 986 '~S001R11 Sealer Ctrlr 2 Required Rezeroing WB2[30].26'; 987 '~S001R11 Mig Barrel Replacement Warning WB2[30].27'; 988 '~S001R11 Mig Barrel Replacement Required WB2[30].28'; 989 '~S001R11 In Touch Up Mode WB2[30].29'; 990 '~S001R11 Touch Up Mode Not Enabled WB2[30].30'; 991 '~Spare WB2[30].31'; 992 '~S001R11 Laser Controller Fault WB2[31].0'; 993 '~S001R11 Laser Dirty Glass Warning WB2[31].1'; 994 '~S001R11 Laser Warning WB2[31].2'; 995 '~Spare WB2[31].3'; 996 '~Spare WB2[31].4'; 997 '~Spare WB2[31].5'; 998 '~Spare WB2[31].6'; 999 '~Spare WB2[31].7'; 1000 '~Spare WB2[31].8'; 1001 '~Spare WB2[31].9'; 1002 '~Spare WB2[31].10'; 1003 '~Spare WB2[31].11'; 1004 '~Spare WB2[31].12'; 1005 '~Spare WB2[31].13'; 1006 '~Spare WB2[31].14'; 1007 '~Spare WB2[31].15'; 1008 '~Spare WB2[31].16'; 1009 '~Spare WB2[31].17'; 1010 '~Spare WB2[31].18'; 1011 '~Spare WB2[31].19'; 1012 '~Spare WB2[31].20'; 1013 '~Spare WB2[31].21'; 1014 '~Spare WB2[31].22'; 1015 '~Spare WB2[31].23'; 1016 '~Spare WB2[31].24'; 1017 '~Spare WB2[31].25'; 1018 '~Spare WB2[31].26'; 1019 '~Spare WB2[31].27'; 1020 '~Spare WB2[31].28'; 1021 '~Spare WB2[31].29'; 1022 '~Spare WB2[31].30'; 1023 '~Spare WB2[31].31'; 1024 '~Spare WB2[32].0'; 1025 '~Spare WB2[32].1'; 1026 '~Spare WB2[32].2'; 1027 '~Spare WB2[32].3'; 1028 '~Spare WB2[32].4'; 1029 '~Spare WB2[32].5'; 1030 '~Spare WB2[32].6'; 1031 '~Spare WB2[32].7'; 1032 '~Spare WB2[32].8'; 1033 '~Spare WB2[32].9'; 1034 '~Spare WB2[32].10'; 1035 '~Spare WB2[32].11'; 1036 '~Spare WB2[32].12'; 1037 '~Spare WB2[32].13'; 1038 '~Spare WB2[32].14'; 1039 '~Spare WB2[32].15'; 1040 '~Spare WB2[32].16'; 1041 '~Spare WB2[32].17'; 1042 '~Spare WB2[32].18'; 1043 '~Spare WB2[32].19'; 1044 '~Spare WB2[32].20'; 1045 '~Spare WB2[32].21'; 1046 '~Spare WB2[32].22'; 1047 '~Spare WB2[32].23'; 1048 '~Spare WB2[32].24'; 1049 '~Spare WB2[32].25'; 1050 '~Spare WB2[32].26'; 1051 '~Spare WB2[32].27'; 1052 '~Spare WB2[32].28'; 1053 '~Spare WB2[32].29'; 1054 '~Spare WB2[32].30'; 1055 '~Spare WB2[32].31'; 1056 '~Spare WB2[33].0'; 1057 '~Spare WB2[33].1'; 1058 '~Spare WB2[33].2'; 1059 '~Spare WB2[33].3'; 1060 '~Spare WB2[33].4'; 1061 '~Spare WB2[33].5'; 1062 '~Spare WB2[33].6'; 1063 '~Spare WB2[33].7'; 1064 '~Spare WB2[33].8'; 1065 '~Spare WB2[33].9'; 1066 '~Spare WB2[33].10'; 1067 '~Spare WB2[33].11'; 1068 '~Spare WB2[33].12'; 1069 '~Spare WB2[33].13'; 1070 '~Spare WB2[33].14'; 1071 '~Spare WB2[33].15'; 1072 '~Spare WB2[33].16'; 1073 '~Spare WB2[33].17'; 1074 '~Spare WB2[33].18'; 1075 '~Spare WB2[33].19'; 1076 '~Spare WB2[33].20'; 1077 '~Spare WB2[33].21'; 1078 '~Spare WB2[33].22'; 1079 '~Spare WB2[33].23'; 1080 '~Spare WB2[33].24'; 1081 '~Spare WB2[33].25'; 1082 '~Spare WB2[33].26'; 1083 '~Spare WB2[33].27'; 1084 '~Spare WB2[33].28'; 1085 '~Spare WB2[33].29'; 1086 '~Spare WB2[33].30'; 1087 '~Spare WB2[33].31'; 1088 '~S001R12 Waiting Zone #1 Not Clear WB2[34].0'; 1089 '~S001R12 Waiting Zone #2 Not Clear WB2[34].1'; 1090 '~S001R12 Waiting Zone #3 Not Clear WB2[34].2'; 1091 '~S001R12 Waiting Zone #4 Not Clear WB2[34].3'; 1092 '~S001R12 Waiting Zone #5 Not Clear WB2[34].4'; 1093 '~S001R12 Waiting Zone #6 Not Clear WB2[34].5'; 1094 '~S001R12 Waiting Zone #7 Not Clear WB2[34].6'; 1095 '~S001R12 Waiting Zone #8 Not Clear WB2[34].7'; 1096 '~S001R12 Waiting Zone #9 Not Clear WB2[34].8'; 1097 '~S001R12 Waiting Zone #10 Not Clear WB2[34].9'; 1098 '~S001R12 Waiting Zone #11 Not Clear WB2[34].10'; 1099 '~S001R12 Waiting Zone #12 Not Clear WB2[34].11'; 1100 '~S001R12 Waiting Zone #13 Not Clear WB2[34].12'; 1101 '~S001R12 Waiting Zone #14 Not Clear WB2[34].13'; 1102 '~S001R12 Waiting Tip Dress Zone #1 Not Clear WB2[34].14'; 1103 '~S001R12 Waiting Tip Dress Zone #2 Not Clear WB2[34].15'; 1104 '~S001R12 Adjacent Robot xx-xx In Teach WB2[34].16'; 1105 '~S001R12 Adjacent Robot xx-xx In Teach WB2[34].17'; 1106 '~S001R12 Adjacent Robot xx-xx In Teach WB2[34].18'; 1107 '~S001R12 Adjacent Robot xx-xx In Teach WB2[34].19'; 1108 '~S001R12 Adjacent Robot xx-xx In Teach WB2[34].20'; 1109 '~S001R12 Adjacent Robot xx-xx In Teach WB2[34].21'; 1110 '~S001R12 Adjacent Robot xx-xx In Teach WB2[34].22'; 1111 '~S001R12 Adjacent Robot xx-xx In Teach WB2[34].23'; 1112 '~S001R12 Adjacent Robot xx-xx In Teach WB2[34].24'; 1113 '~S001R12 Adjacent Robot xx-xx In Teach WB2[34].25'; 1114 '~Spare WB2[34].26'; 1115 '~Spare WB2[34].27'; 1116 '~Spare WB2[34].28'; 1117 '~S001R12 Robot Not Clear Of Fixture WB2[34].29'; 1118 '~Spare WB2[34].30'; 1119 '~Spare WB2[34].31'; 1120 '~Spare WB2[35].0'; 1121 '~Spare WB2[35].1'; 1122 '~Spare WB2[35].2'; 1123 '~Spare WB2[35].3'; 1124 '~Spare WB2[35].4'; 1125 '~Spare WB2[35].5'; 1126 '~Spare WB2[35].6'; 1127 '~Spare WB2[35].7'; 1128 '~Spare WB2[35].8'; 1129 '~Spare WB2[35].9'; 1130 '~Spare WB2[35].10'; 1131 '~Spare WB2[35].11'; 1132 '~Spare WB2[35].12'; 1133 '~Spare WB2[35].13'; 1134 '~Spare WB2[35].14'; 1135 '~Spare WB2[35].15'; 1136 '~Spare WB2[35].16'; 1137 '~Spare WB2[35].17'; 1138 '~Spare WB2[35].18'; 1139 '~Spare WB2[35].19'; 1140 '~Spare WB2[35].20'; 1141 '~Spare WB2[35].21'; 1142 '~Spare WB2[35].22'; 1143 '~Spare WB2[35].23'; 1144 '~Spare WB2[35].24'; 1145 '~Spare WB2[35].25'; 1146 '~Spare WB2[35].26'; 1147 '~Spare WB2[35].27'; 1148 '~Spare WB2[35].28'; 1149 '~Spare WB2[35].29'; 1150 '~Spare WB2[35].30'; 1151 '~Spare WB2[35].31'; 1152 '~S001R12 Cycle Overtime WB2[36].0'; 1153 '~S001R12 In Bypass WB2[36].1'; 1154 '~S001R12 Battery Low WB2[36].2'; 1155 '~S001R12 Servo Over Torque WB2[36].3'; 1156 '~S001R12 Process Retry In Progress WB2[36].4'; 1157 '~Spare WB2[36].5'; 1158 '~S001R12 Robot Edit Occurred Ext App WB2[36].6'; 1159 '~S001R12 Robot Input Simmed WB2[36].7'; 1160 '~S001R12 Robot Output Simmed WB2[36].8'; 1161 '~Spare WB2[36].9'; 1162 '~Spare WB2[36].10'; 1163 '~Spare WB2[36].11'; 1164 '~Spare WB2[36].12'; 1165 '~Spare WB2[36].13'; 1166 '~Spare WB2[36].14'; 1167 '~Spare WB2[36].15'; 1168 '~S001R12F1B1.M.ModuleFlt - Externa App 1 I/O Module Warning WB2[36].16'; 1169 '~S001R12F2B1.M.ModuleFlt - Externa App 2 I/O Module Warning WB2[36].17'; 1170 '~S001R12F3B1.M.ModuleFlt - Externa App 3 I/O Module Warning WB2[36].18'; 1171 '~Spare WB2[36].19'; 1172 '~Spare WB2[36].20'; 1173 '~Spare WB2[36].21'; 1174 '~Spare WB2[36].22'; 1175 '~Spare WB2[36].23'; 1176 '~S001R12ES1 - S001R12 EtherNet Switch Port At Half Duplex WB2[36].24'; 1177 '~S001R12ES1 - S001R12 EtherNet Switch Config Changes Not Saved WB2[36].25'; 1178 '~S001R12ES1 - S001R12 EtherNet Switch Configuration Changed WB2[36].26'; 1179 '~S001R12ES1 - S001R12 EtherNet Switch Port With Excessive Errors WB2[36].27'; 1180 '~S001R12ES1 - S001R12 EtherNet Switch Port With Utilization Warning WB2[36].28'; 1181 '~S001R12ES1 - S001R12 EtherNet Switch Changes Require Reboot WB2[36].29'; 1182 '~Spare WB2[36].30'; 1183 '~Spare WB2[36].31'; 1184 '~Spare WB2[37].0'; 1185 '~Spare WB2[37].1'; 1186 '~S001R12 Servo Gun Tip Calib Request 1 WB2[37].2'; 1187 '~S001R12 I-Available Warning 1 WB2[37].3'; 1188 '~S001R12 Tip Dress Motor 1 Fault Bypassed WB2[37].4'; 1189 '~S001R12 Tip Change Notice 1 WB2[37].5'; 1190 '~S001R12 Bypass Tip Dresser 1 Selected WB2[37].6'; 1191 '~S001R12 Auto Tip Changer Low 1 WB2[37].7'; 1192 '~S001R12 Auto Tip Changer Empty 1 WB2[37].8'; 1193 '~S001R12 Tip Wear Ratio Warning 1 - Touch Up Tip Dress Program WB2[37].9'; 1194 '~S001R12 Stud Weld 1 Maintenance Reqd WB2[37].10'; 1195 '~S001R12 Stud Weld 1 Low Stud Warning WB2[37].11'; 1196 '~Spare WB2[37].12'; 1197 '~S001R12 Rivet 1 Low Rivet Warning WB2[37].13'; 1198 '~S001R12 Rivet 1 - Skip Once Initiated from Robot TP WB2[37].14'; 1199 '~S001R12 Rivet 1 - Skip Remaining Initiated from Robot TP WB2[37].15'; 1200 '~S001R12 Rivet 1 Preventive Maintenace Required WB2[37].16'; 1201 '~S001R12 Rivet 1 Magazine Low WB2[37].17'; 1202 '~S001R12 Tip Change 1 Bypassed WB2[37].18'; 1203 '~S001R12 Mig Weld Fluid Level Low WB2[37].19'; 1204 '~S001R12 Weld Ctrlr 1 Adaptive Mode Is Disabled WB2[37].20'; 1205 '~S001R12 Tip Cutter 1 Warning WB2[37].21'; 1206 '~S001R12 Rivet 1 Tape-Cut Required WB2[37].22'; 1207 '~S001R12 Wire Feeder Motor Over Current WB2[37].23'; 1208 '~Spare WB2[37].24'; 1209 '~S001R12 Sealer Ctrlr 1 Minor Fault WB2[37].25'; 1210 '~S001R12 Sealer Ctrlr 1 Required Rezeroing WB2[37].26'; 1211 '~S001R12 Loaded To Average WB2[37].27'; 1212 '~S001R12 Vision Process Aborted WB2[37].28'; 1213 '~S001R12 Vision System Trending WB2[37].29'; 1214 '~S001R12 Vision Out Of Tolerance WB2[37].30'; 1215 '~Spare WB2[37].31'; 1216 '~Spare WB2[38].0'; 1217 '~Spare WB2[38].1'; 1218 '~S001R12 Servo Gun Tip Calib Request 2 WB2[38].2'; 1219 '~S001R12 I-Available Warning 2 WB2[38].3'; 1220 '~S001R12 Tip Dress Motor 2 Fault Bypassed WB2[38].4'; 1221 '~S001R12 Tip Change Notice 2 WB2[38].5'; 1222 '~S001R12 Bypass Tip Dresser 2 Selected WB2[38].6'; 1223 '~S001R12 Auto Tip Changer Low 2 WB2[38].7'; 1224 '~S001R12 Auto Tip Changer Empty 2 WB2[38].8'; 1225 '~S001R12 Tip Wear Ratio Warning 2 - Touch Up Tip Dress Program WB2[38].9'; 1226 '~S001R12 Stud Weld 2 Maintenance Reqd WB2[38].10'; 1227 '~S001R12 Stud Weld 2 Low Stud Warning WB2[38].11'; 1228 '~Spare WB2[38].12'; 1229 '~S001R12 Rivet 2 Low Rivet Warning WB2[38].13'; 1230 '~S001R12 Rivet 2 - Skip Once Initiated from Robot TP WB2[38].14'; 1231 '~S001R12 Rivet 2 - Skip Remaining Initiated from Robot TP WB2[38].15'; 1232 '~S001R12 Rivet 2 Preventive Maintenace Required WB2[38].16'; 1233 '~S001R12 Rivet 2 Magazine Low WB2[38].17'; 1234 '~S001R12 Tip Change 2 Bypassed WB2[38].18'; 1235 '~S001R12 Laser Dirty Glass Warning WB2[38].19'; 1236 '~S001R12 Weld Ctrlr 2 Adaptive Mode Is Disabled WB2[38].20'; 1237 '~S001R12 Tip Cutter 2 Warning WB2[38].21'; 1238 '~S001R12 Rivet 2 Tape-Cut Required WB2[38].22'; 1239 '~S001R12 Mig Tip Nozzel Replacement Warning WB2[38].23'; 1240 '~S001R12 Mig Tip Nozzel Replacement Required WB2[38].24'; 1241 '~S001R12 Sealer Ctrlr 2 Minor Fault WB2[38].25'; 1242 '~S001R12 Sealer Ctrlr 2 Required Rezeroing WB2[38].26'; 1243 '~S001R12 Mig Barrel Replacement Warning WB2[38].27'; 1244 '~S001R12 Mig Barrel Replacement Required WB2[38].28'; 1245 '~S001R12 In Touch Up Mode WB2[38].29'; 1246 '~S001R12 Touch Up Mode Not Enabled WB2[38].30'; 1247 '~Spare WB2[38].31'; 1248 '~S001R12 Laser Controller Fault WB2[39].0'; 1249 '~S001R12 Laser Dirty Glass Warning WB2[39].1'; 1250 '~S001R12 Laser Warning WB2[39].2'; 1251 '~Spare WB2[39].3'; 1252 '~Spare WB2[39].4'; 1253 '~Spare WB2[39].5'; 1254 '~Spare WB2[39].6'; 1255 '~Spare WB2[39].7'; 1256 '~Spare WB2[39].8'; 1257 '~Spare WB2[39].9'; 1258 '~Spare WB2[39].10'; 1259 '~Spare WB2[39].11'; 1260 '~Spare WB2[39].12'; 1261 '~Spare WB2[39].13'; 1262 '~Spare WB2[39].14'; 1263 '~Spare WB2[39].15'; 1264 '~Spare WB2[39].16'; 1265 '~Spare WB2[39].17'; 1266 '~Spare WB2[39].18'; 1267 '~Spare WB2[39].19'; 1268 '~Spare WB2[39].20'; 1269 '~Spare WB2[39].21'; 1270 '~Spare WB2[39].22'; 1271 '~Spare WB2[39].23'; 1272 '~Spare WB2[39].24'; 1273 '~Spare WB2[39].25'; 1274 '~Spare WB2[39].26'; 1275 '~Spare WB2[39].27'; 1276 '~Spare WB2[39].28'; 1277 '~Spare WB2[39].29'; 1278 '~Spare WB2[39].30'; 1279 '~Spare WB2[39].31'; 1280 '~Spare WB2[40].0'; 1281 '~Spare WB2[40].1'; 1282 '~Spare WB2[40].2'; 1283 '~Spare WB2[40].3'; 1284 '~Spare WB2[40].4'; 1285 '~Spare WB2[40].5'; 1286 '~Spare WB2[40].6'; 1287 '~Spare WB2[40].7'; 1288 '~Spare WB2[40].8'; 1289 '~Spare WB2[40].9'; 1290 '~Spare WB2[40].10'; 1291 '~Spare WB2[40].11'; 1292 '~Spare WB2[40].12'; 1293 '~Spare WB2[40].13'; 1294 '~Spare WB2[40].14'; 1295 '~Spare WB2[40].15'; 1296 '~Spare WB2[40].16'; 1297 '~Spare WB2[40].17'; 1298 '~Spare WB2[40].18'; 1299 '~Spare WB2[40].19'; 1300 '~Spare WB2[40].20'; 1301 '~Spare WB2[40].21'; 1302 '~Spare WB2[40].22'; 1303 '~Spare WB2[40].23'; 1304 '~Spare WB2[40].24'; 1305 '~Spare WB2[40].25'; 1306 '~Spare WB2[40].26'; 1307 '~Spare WB2[40].27'; 1308 '~Spare WB2[40].28'; 1309 '~Spare WB2[40].29'; 1310 '~Spare WB2[40].30'; 1311 '~Spare WB2[40].31'; 1312 '~Spare WB2[41].0'; 1313 '~Spare WB2[41].1'; 1314 '~Spare WB2[41].2'; 1315 '~Spare WB2[41].3'; 1316 '~Spare WB2[41].4'; 1317 '~Spare WB2[41].5'; 1318 '~Spare WB2[41].6'; 1319 '~Spare WB2[41].7'; 1320 '~Spare WB2[41].8'; 1321 '~Spare WB2[41].9'; 1322 '~Spare WB2[41].10'; 1323 '~Spare WB2[41].11'; 1324 '~Spare WB2[41].12'; 1325 '~Spare WB2[41].13'; 1326 '~Spare WB2[41].14'; 1327 '~Spare WB2[41].15'; 1328 '~Spare WB2[41].16'; 1329 '~Spare WB2[41].17'; 1330 '~Spare WB2[41].18'; 1331 '~Spare WB2[41].19'; 1332 '~Spare WB2[41].20'; 1333 '~Spare WB2[41].21'; 1334 '~Spare WB2[41].22'; 1335 '~Spare WB2[41].23'; 1336 '~Spare WB2[41].24'; 1337 '~Spare WB2[41].25'; 1338 '~Spare WB2[41].26'; 1339 '~Spare WB2[41].27'; 1340 '~Spare WB2[41].28'; 1341 '~Spare WB2[41].29'; 1342 '~Spare WB2[41].30'; 1343 '~Spare WB2[41].31'; 1344 '~S001R13 Waiting Zone #1 Not Clear WB2[42].0'; 1345 '~S001R13 Waiting Zone #2 Not Clear WB2[42].1'; 1346 '~S001R13 Waiting Zone #3 Not Clear WB2[42].2'; 1347 '~S001R13 Waiting Zone #4 Not Clear WB2[42].3'; 1348 '~S001R13 Waiting Zone #5 Not Clear WB2[42].4'; 1349 '~S001R13 Waiting Zone #6 Not Clear WB2[42].5'; 1350 '~S001R13 Waiting Zone #7 Not Clear WB2[42].6'; 1351 '~S001R13 Waiting Zone #8 Not Clear WB2[42].7'; 1352 '~S001R13 Waiting Zone #9 Not Clear WB2[42].8'; 1353 '~S001R13 Waiting Zone #10 Not Clear WB2[42].9'; 1354 '~S001R13 Waiting Zone #11 Not Clear WB2[42].10'; 1355 '~S001R13 Waiting Zone #12 Not Clear WB2[42].11'; 1356 '~S001R13 Waiting Zone #13 Not Clear WB2[42].12'; 1357 '~S001R13 Waiting Zone #14 Not Clear WB2[42].13'; 1358 '~S001R13 Waiting Tip Dress Zone #1 Not Clear WB2[42].14'; 1359 '~S001R13 Waiting Tip Dress Zone #2 Not Clear WB2[42].15'; 1360 '~S001R13 Adjacent Robot xx-xx In Teach WB2[42].16'; 1361 '~S001R13 Adjacent Robot xx-xx In Teach WB2[42].17'; 1362 '~S001R13 Adjacent Robot xx-xx In Teach WB2[42].18'; 1363 '~S001R13 Adjacent Robot xx-xx In Teach WB2[42].19'; 1364 '~S001R13 Adjacent Robot xx-xx In Teach WB2[42].20'; 1365 '~S001R13 Adjacent Robot xx-xx In Teach WB2[42].21'; 1366 '~S001R13 Adjacent Robot xx-xx In Teach WB2[42].22'; 1367 '~S001R13 Adjacent Robot xx-xx In Teach WB2[42].23'; 1368 '~S001R13 Adjacent Robot xx-xx In Teach WB2[42].24'; 1369 '~S001R13 Adjacent Robot xx-xx In Teach WB2[42].25'; 1370 '~Spare WB2[42].26'; 1371 '~Spare WB2[42].27'; 1372 '~Spare WB2[42].28'; 1373 '~S001R13 Robot Not Clear Of Fixture WB2[42].29'; 1374 '~Spare WB2[42].30'; 1375 '~Spare WB2[42].31'; 1376 '~Spare WB2[43].0'; 1377 '~Spare WB2[43].1'; 1378 '~Spare WB2[43].2'; 1379 '~Spare WB2[43].3'; 1380 '~Spare WB2[43].4'; 1381 '~Spare WB2[43].5'; 1382 '~Spare WB2[43].6'; 1383 '~Spare WB2[43].7'; 1384 '~Spare WB2[43].8'; 1385 '~Spare WB2[43].9'; 1386 '~Spare WB2[43].10'; 1387 '~Spare WB2[43].11'; 1388 '~Spare WB2[43].12'; 1389 '~Spare WB2[43].13'; 1390 '~Spare WB2[43].14'; 1391 '~Spare WB2[43].15'; 1392 '~Spare WB2[43].16'; 1393 '~Spare WB2[43].17'; 1394 '~Spare WB2[43].18'; 1395 '~Spare WB2[43].19'; 1396 '~Spare WB2[43].20'; 1397 '~Spare WB2[43].21'; 1398 '~Spare WB2[43].22'; 1399 '~Spare WB2[43].23'; 1400 '~Spare WB2[43].24'; 1401 '~Spare WB2[43].25'; 1402 '~Spare WB2[43].26'; 1403 '~Spare WB2[43].27'; 1404 '~Spare WB2[43].28'; 1405 '~Spare WB2[43].29'; 1406 '~Spare WB2[43].30'; 1407 '~Spare WB2[43].31'; 1408 '~S001R13 Cycle Overtime WB2[44].0'; 1409 '~S001R13 In Bypass WB2[44].1'; 1410 '~S001R13 Battery Low WB2[44].2'; 1411 '~S001R13 Servo Over Torque WB2[44].3'; 1412 '~S001R13 Process Retry In Progress WB2[44].4'; 1413 '~Spare WB2[44].5'; 1414 '~S001R13 Robot Edit Occurred Ext App WB2[44].6'; 1415 '~S001R13 Robot Input Simmed WB2[44].7'; 1416 '~S001R13 Robot Output Simmed WB2[44].8'; 1417 '~Spare WB2[44].9'; 1418 '~Spare WB2[44].10'; 1419 '~Spare WB2[44].11'; 1420 '~Spare WB2[44].12'; 1421 '~Spare WB2[44].13'; 1422 '~Spare WB2[44].14'; 1423 '~Spare WB2[44].15'; 1424 '~S001R13F1B1.M.ModuleFlt - Externa App 1 I/O Module Warning WB2[44].16'; 1425 '~S001R13F2B1.M.ModuleFlt - Externa App 2 I/O Module Warning WB2[44].17'; 1426 '~S001R13F3B1.M.ModuleFlt - Externa App 3 I/O Module Warning WB2[44].18'; 1427 '~Spare WB2[44].19'; 1428 '~Spare WB2[44].20'; 1429 '~Spare WB2[44].21'; 1430 '~Spare WB2[44].22'; 1431 '~Spare WB2[44].23'; 1432 '~S001R13ES1 - S001R13 EtherNet Switch Port At Half Duplex WB2[44].24'; 1433 '~S001R13ES1 - S001R13 EtherNet Switch Config Changes Not Saved WB2[44].25'; 1434 '~S001R13ES1 - S001R13 EtherNet Switch Configuration Changed WB2[44].26'; 1435 '~S001R13ES1 - S001R13 EtherNet Switch Port With Excessive Errors WB2[44].27'; 1436 '~S001R13ES1 - S001R13 EtherNet Switch Port With Utilization Warning WB2[44].28'; 1437 '~S001R13ES1 - S001R13 EtherNet Switch Changes Require Reboot WB2[44].29'; 1438 '~Spare WB2[44].30'; 1439 '~Spare WB2[44].31'; 1440 '~Spare WB2[45].0'; 1441 '~Spare WB2[45].1'; 1442 '~S001R13 Servo Gun Tip Calib Request 1 WB2[45].2'; 1443 '~S001R13 I-Available Warning 1 WB2[45].3'; 1444 '~S001R13 Tip Dress Motor 1 Fault Bypassed WB2[45].4'; 1445 '~S001R13 Tip Change Notice 1 WB2[45].5'; 1446 '~S001R13 Bypass Tip Dresser 1 Selected WB2[45].6'; 1447 '~S001R13 Auto Tip Changer Low 1 WB2[45].7'; 1448 '~S001R13 Auto Tip Changer Empty 1 WB2[45].8'; 1449 '~S001R13 Tip Wear Ratio Warning 1 - Touch Up Tip Dress Program WB2[45].9'; 1450 '~S001R13 Stud Weld 1 Maintenance Reqd WB2[45].10'; 1451 '~S001R13 Stud Weld 1 Low Stud Warning WB2[45].11'; 1452 '~Spare WB2[45].12'; 1453 '~S001R13 Rivet 1 Low Rivet Warning WB2[45].13'; 1454 '~S001R13 Rivet 1 - Skip Once Initiated from Robot TP WB2[45].14'; 1455 '~S001R13 Rivet 1 - Skip Remaining Initiated from Robot TP WB2[45].15'; 1456 '~S001R13 Rivet 1 Preventive Maintenace Required WB2[45].16'; 1457 '~S001R13 Rivet 1 Magazine Low WB2[45].17'; 1458 '~S001R13 Tip Change 1 Bypassed WB2[45].18'; 1459 '~S001R13 Mig Weld Fluid Level Low WB2[45].19'; 1460 '~S001R13 Weld Ctrlr 1 Adaptive Mode Is Disabled WB2[45].20'; 1461 '~S001R13 Tip Cutter 1 Warning WB2[45].21'; 1462 '~S001R13 Rivet 1 Tape-Cut Required WB2[45].22'; 1463 '~S001R13 Wire Feeder Motor Over Current WB2[45].23'; 1464 '~Spare WB2[45].24'; 1465 '~S001R13 Sealer Ctrlr 1 Minor Fault WB2[45].25'; 1466 '~S001R13 Sealer Ctrlr 1 Required Rezeroing WB2[45].26'; 1467 '~S001R13 Loaded To Average WB2[45].27'; 1468 '~S001R13 Vision Process Aborted WB2[45].28'; 1469 '~S001R13 Vision System Trending WB2[45].29'; 1470 '~S001R13 Vision Out Of Tolerance WB2[45].30'; 1471 '~Spare WB2[45].31'; 1472 '~Spare WB2[46].0'; 1473 '~Spare WB2[46].1'; 1474 '~S001R13 Servo Gun Tip Calib Request 2 WB2[46].2'; 1475 '~S001R13 I-Available Warning 2 WB2[46].3'; 1476 '~S001R13 Tip Dress Motor 2 Fault Bypassed WB2[46].4'; 1477 '~S001R13 Tip Change Notice 2 WB2[46].5'; 1478 '~S001R13 Bypass Tip Dresser 2 Selected WB2[46].6'; 1479 '~S001R13 Auto Tip Changer Low 2 WB2[46].7'; 1480 '~S001R13 Auto Tip Changer Empty 2 WB2[46].8'; 1481 '~S001R13 Tip Wear Ratio Warning 2 - Touch Up Tip Dress Program WB2[46].9'; 1482 '~S001R13 Stud Weld 2 Maintenance Reqd WB2[46].10'; 1483 '~S001R13 Stud Weld 2 Low Stud Warning WB2[46].11'; 1484 '~Spare WB2[46].12'; 1485 '~S001R13 Rivet 2 Low Rivet Warning WB2[46].13'; 1486 '~S001R13 Rivet 2 - Skip Once Initiated from Robot TP WB2[46].14'; 1487 '~S001R13 Rivet 2 - Skip Remaining Initiated from Robot TP WB2[46].15'; 1488 '~S001R13 Rivet 2 Preventive Maintenace Required WB2[46].16'; 1489 '~S001R13 Rivet 2 Magazine Low WB2[46].17'; 1490 '~S001R13 Tip Change 2 Bypassed WB2[46].18'; 1491 '~S001R13 Laser Dirty Glass Warning WB2[46].19'; 1492 '~S001R13 Weld Ctrlr 2 Adaptive Mode Is Disabled WB2[46].20'; 1493 '~S001R13 Tip Cutter 2 Warning WB2[46].21'; 1494 '~S001R13 Rivet 2 Tape-Cut Required WB2[46].22'; 1495 '~S001R13 Mig Tip Nozzel Replacement Warning WB2[46].23'; 1496 '~S001R13 Mig Tip Nozzel Replacement Required WB2[46].24'; 1497 '~S001R13 Sealer Ctrlr 2 Minor Fault WB2[46].25'; 1498 '~S001R13 Sealer Ctrlr 2 Required Rezeroing WB2[46].26'; 1499 '~S001R13 Mig Barrel Replacement Warning WB2[46].27'; 1500 '~S001R13 Mig Barrel Replacement Required WB2[46].28'; 1501 '~S001R13 In Touch Up Mode WB2[46].29'; 1502 '~S001R13 Touch Up Mode Not Enabled WB2[46].30'; 1503 '~Spare WB2[46].31'; 1504 '~S001R13 Laser Controller Fault WB2[47].0'; 1505 '~S001R13 Laser Dirty Glass Warning WB2[47].1'; 1506 '~S001R13 Laser Warning WB2[47].2'; 1507 '~Spare WB2[47].3'; 1508 '~Spare WB2[47].4'; 1509 '~Spare WB2[47].5'; 1510 '~Spare WB2[47].6'; 1511 '~Spare WB2[47].7'; 1512 '~Spare WB2[47].8'; 1513 '~Spare WB2[47].9'; 1514 '~Spare WB2[47].10'; 1515 '~Spare WB2[47].11'; 1516 '~Spare WB2[47].12'; 1517 '~Spare WB2[47].13'; 1518 '~Spare WB2[47].14'; 1519 '~Spare WB2[47].15'; 1520 '~Spare WB2[47].16'; 1521 '~Spare WB2[47].17'; 1522 '~Spare WB2[47].18'; 1523 '~Spare WB2[47].19'; 1524 '~Spare WB2[47].20'; 1525 '~Spare WB2[47].21'; 1526 '~Spare WB2[47].22'; 1527 '~Spare WB2[47].23'; 1528 '~Spare WB2[47].24'; 1529 '~Spare WB2[47].25'; 1530 '~Spare WB2[47].26'; 1531 '~Spare WB2[47].27'; 1532 '~Spare WB2[47].28'; 1533 '~Spare WB2[47].29'; 1534 '~Spare WB2[47].30'; 1535 '~Spare WB2[47].31'; 1536 '~Spare WB2[48].0'; 1537 '~Spare WB2[48].1'; 1538 '~Spare WB2[48].2'; 1539 '~Spare WB2[48].3'; 1540 '~Spare WB2[48].4'; 1541 '~Spare WB2[48].5'; 1542 '~Spare WB2[48].6'; 1543 '~Spare WB2[48].7'; 1544 '~Spare WB2[48].8'; 1545 '~Spare WB2[48].9'; 1546 '~Spare WB2[48].10'; 1547 '~Spare WB2[48].11'; 1548 '~Spare WB2[48].12'; 1549 '~Spare WB2[48].13'; 1550 '~Spare WB2[48].14'; 1551 '~Spare WB2[48].15'; 1552 '~Spare WB2[48].16'; 1553 '~Spare WB2[48].17'; 1554 '~Spare WB2[48].18'; 1555 '~Spare WB2[48].19'; 1556 '~Spare WB2[48].20'; 1557 '~Spare WB2[48].21'; 1558 '~Spare WB2[48].22'; 1559 '~Spare WB2[48].23'; 1560 '~Spare WB2[48].24'; 1561 '~Spare WB2[48].25'; 1562 '~Spare WB2[48].26'; 1563 '~Spare WB2[48].27'; 1564 '~Spare WB2[48].28'; 1565 '~Spare WB2[48].29'; 1566 '~Spare WB2[48].30'; 1567 '~Spare WB2[48].31'; 1568 '~Spare WB2[49].0'; 1569 '~Spare WB2[49].1'; 1570 '~Spare WB2[49].2'; 1571 '~Spare WB2[49].3'; 1572 '~Spare WB2[49].4'; 1573 '~Spare WB2[49].5'; 1574 '~Spare WB2[49].6'; 1575 '~Spare WB2[49].7'; 1576 '~Spare WB2[49].8'; 1577 '~Spare WB2[49].9'; 1578 '~Spare WB2[49].10'; 1579 '~Spare WB2[49].11'; 1580 '~Spare WB2[49].12'; 1581 '~Spare WB2[49].13'; 1582 '~Spare WB2[49].14'; 1583 '~Spare WB2[49].15'; 1584 '~Spare WB2[49].16'; 1585 '~Spare WB2[49].17'; 1586 '~Spare WB2[49].18'; 1587 '~Spare WB2[49].19'; 1588 '~Spare WB2[49].20'; 1589 '~Spare WB2[49].21'; 1590 '~Spare WB2[49].22'; 1591 '~Spare WB2[49].23'; 1592 '~Spare WB2[49].24'; 1593 '~Spare WB2[49].25'; 1594 '~Spare WB2[49].26'; 1595 '~Spare WB2[49].27'; 1596 '~Spare WB2[49].28'; 1597 '~Spare WB2[49].29'; 1598 '~Spare WB2[49].30'; 1599 '~Spare WB2[49].31'; 1600 '~S001R14 Waiting Zone #1 Not Clear WB2[50].0'; 1601 '~S001R14 Waiting Zone #2 Not Clear WB2[50].1'; 1602 '~S001R14 Waiting Zone #3 Not Clear WB2[50].2'; 1603 '~S001R14 Waiting Zone #4 Not Clear WB2[50].3'; 1604 '~S001R14 Waiting Zone #5 Not Clear WB2[50].4'; 1605 '~S001R14 Waiting Zone #6 Not Clear WB2[50].5'; 1606 '~S001R14 Waiting Zone #7 Not Clear WB2[50].6'; 1607 '~S001R14 Waiting Zone #8 Not Clear WB2[50].7'; 1608 '~S001R14 Waiting Zone #9 Not Clear WB2[50].8'; 1609 '~S001R14 Waiting Zone #10 Not Clear WB2[50].9'; 1610 '~S001R14 Waiting Zone #11 Not Clear WB2[50].10'; 1611 '~S001R14 Waiting Zone #12 Not Clear WB2[50].11'; 1612 '~S001R14 Waiting Zone #13 Not Clear WB2[50].12'; 1613 '~S001R14 Waiting Zone #14 Not Clear WB2[50].13'; 1614 '~S001R14 Waiting Tip Dress Zone #1 Not Clear WB2[50].14'; 1615 '~S001R14 Waiting Tip Dress Zone #2 Not Clear WB2[50].15'; 1616 '~S001R14 Adjacent Robot xx-xx In Teach WB2[50].16'; 1617 '~S001R14 Adjacent Robot xx-xx In Teach WB2[50].17'; 1618 '~S001R14 Adjacent Robot xx-xx In Teach WB2[50].18'; 1619 '~S001R14 Adjacent Robot xx-xx In Teach WB2[50].19'; 1620 '~S001R14 Adjacent Robot xx-xx In Teach WB2[50].20'; 1621 '~S001R14 Adjacent Robot xx-xx In Teach WB2[50].21'; 1622 '~S001R14 Adjacent Robot xx-xx In Teach WB2[50].22'; 1623 '~S001R14 Adjacent Robot xx-xx In Teach WB2[50].23'; 1624 '~S001R14 Adjacent Robot xx-xx In Teach WB2[50].24'; 1625 '~S001R14 Adjacent Robot xx-xx In Teach WB2[50].25'; 1626 '~Spare WB2[50].26'; 1627 '~Spare WB2[50].27'; 1628 '~Spare WB2[50].28'; 1629 '~S001R14 Robot Not Clear Of Fixture WB2[50].29'; 1630 '~Spare WB2[50].30'; 1631 '~Spare WB2[50].31'; 1632 '~Spare WB2[51].0'; 1633 '~Spare WB2[51].1'; 1634 '~Spare WB2[51].2'; 1635 '~Spare WB2[51].3'; 1636 '~Spare WB2[51].4'; 1637 '~Spare WB2[51].5'; 1638 '~Spare WB2[51].6'; 1639 '~Spare WB2[51].7'; 1640 '~Spare WB2[51].8'; 1641 '~Spare WB2[51].9'; 1642 '~Spare WB2[51].10'; 1643 '~Spare WB2[51].11'; 1644 '~Spare WB2[51].12'; 1645 '~Spare WB2[51].13'; 1646 '~Spare WB2[51].14'; 1647 '~Spare WB2[51].15'; 1648 '~Spare WB2[51].16'; 1649 '~Spare WB2[51].17'; 1650 '~Spare WB2[51].18'; 1651 '~Spare WB2[51].19'; 1652 '~Spare WB2[51].20'; 1653 '~Spare WB2[51].21'; 1654 '~Spare WB2[51].22'; 1655 '~Spare WB2[51].23'; 1656 '~Spare WB2[51].24'; 1657 '~Spare WB2[51].25'; 1658 '~Spare WB2[51].26'; 1659 '~Spare WB2[51].27'; 1660 '~Spare WB2[51].28'; 1661 '~Spare WB2[51].29'; 1662 '~Spare WB2[51].30'; 1663 '~Spare WB2[51].31'; 1664 '~S001R14 Cycle Overtime WB2[52].0'; 1665 '~S001R14 In Bypass WB2[52].1'; 1666 '~S001R14 Battery Low WB2[52].2'; 1667 '~S001R14 Servo Over Torque WB2[52].3'; 1668 '~S001R14 Process Retry In Progress WB2[52].4'; 1669 '~Spare WB2[52].5'; 1670 '~S001R14 Robot Edit Occurred Ext App WB2[52].6'; 1671 '~S001R14 Robot Input Simmed WB2[52].7'; 1672 '~S001R14 Robot Output Simmed WB2[52].8'; 1673 '~Spare WB2[52].9'; 1674 '~Spare WB2[52].10'; 1675 '~Spare WB2[52].11'; 1676 '~Spare WB2[52].12'; 1677 '~Spare WB2[52].13'; 1678 '~Spare WB2[52].14'; 1679 '~Spare WB2[52].15'; 1680 '~S001R14F1B1.M.ModuleFlt - Externa App 1 I/O Module Warning WB2[52].16'; 1681 '~S001R14F2B1.M.ModuleFlt - Externa App 2 I/O Module Warning WB2[52].17'; 1682 '~S001R14F3B1.M.ModuleFlt - Externa App 3 I/O Module Warning WB2[52].18'; 1683 '~Spare WB2[52].19'; 1684 '~Spare WB2[52].20'; 1685 '~Spare WB2[52].21'; 1686 '~Spare WB2[52].22'; 1687 '~Spare WB2[52].23'; 1688 '~S001R14ES1 - S001R14 EtherNet Switch Port At Half Duplex WB2[52].24'; 1689 '~S001R14ES1 - S001R14 EtherNet Switch Config Changes Not Saved WB2[52].25'; 1690 '~S001R14ES1 - S001R14 EtherNet Switch Configuration Changed WB2[52].26'; 1691 '~S001R14ES1 - S001R14 EtherNet Switch Port With Excessive Errors WB2[52].27'; 1692 '~S001R14ES1 - S001R14 EtherNet Switch Port With Utilization Warning WB2[52].28'; 1693 '~S001R14ES1 - S001R14 EtherNet Switch Changes Require Reboot WB2[52].29'; 1694 '~Spare WB2[52].30'; 1695 '~Spare WB2[52].31'; 1696 '~Spare WB2[53].0'; 1697 '~Spare WB2[53].1'; 1698 '~S001R14 Servo Gun Tip Calib Request 1 WB2[53].2'; 1699 '~S001R14 I-Available Warning 1 WB2[53].3'; 1700 '~S001R14 Tip Dress Motor 1 Fault Bypassed WB2[53].4'; 1701 '~S001R14 Tip Change Notice 1 WB2[53].5'; 1702 '~S001R14 Bypass Tip Dresser 1 Selected WB2[53].6'; 1703 '~S001R14 Auto Tip Changer Low 1 WB2[53].7'; 1704 '~S001R14 Auto Tip Changer Empty 1 WB2[53].8'; 1705 '~S001R14 Tip Wear Ratio Warning 1 - Touch Up Tip Dress Program WB2[53].9'; 1706 '~S001R14 Stud Weld 1 Maintenance Reqd WB2[53].10'; 1707 '~S001R14 Stud Weld 1 Low Stud Warning WB2[53].11'; 1708 '~Spare WB2[53].12'; 1709 '~S001R14 Rivet 1 Low Rivet Warning WB2[53].13'; 1710 '~S001R14 Rivet 1 - Skip Once Initiated from Robot TP WB2[53].14'; 1711 '~S001R14 Rivet 1 - Skip Remaining Initiated from Robot TP WB2[53].15'; 1712 '~S001R14 Rivet 1 Preventive Maintenace Required WB2[53].16'; 1713 '~S001R14 Rivet 1 Magazine Low WB2[53].17'; 1714 '~S001R14 Tip Change 1 Bypassed WB2[53].18'; 1715 '~S001R14 Mig Weld Fluid Level Low WB2[53].19'; 1716 '~S001R14 Weld Ctrlr 1 Adaptive Mode Is Disabled WB2[53].20'; 1717 '~S001R14 Tip Cutter 1 Warning WB2[53].21'; 1718 '~S001R14 Rivet 1 Tape-Cut Required WB2[53].22'; 1719 '~S001R14 Wire Feeder Motor Over Current WB2[53].23'; 1720 '~Spare WB2[53].24'; 1721 '~S001R14 Sealer Ctrlr 1 Minor Fault WB2[53].25'; 1722 '~S001R14 Sealer Ctrlr 1 Required Rezeroing WB2[53].26'; 1723 '~S001R14 Loaded To Average WB2[53].27'; 1724 '~S001R14 Vision Process Aborted WB2[53].28'; 1725 '~S001R14 Vision System Trending WB2[53].29'; 1726 '~S001R14 Vision Out Of Tolerance WB2[53].30'; 1727 '~Spare WB2[53].31'; 1728 '~Spare WB2[54].0'; 1729 '~Spare WB2[54].1'; 1730 '~S001R14 Servo Gun Tip Calib Request 2 WB2[54].2'; 1731 '~S001R14 I-Available Warning 2 WB2[54].3'; 1732 '~S001R14 Tip Dress Motor 2 Fault Bypassed WB2[54].4'; 1733 '~S001R14 Tip Change Notice 2 WB2[54].5'; 1734 '~S001R14 Bypass Tip Dresser 2 Selected WB2[54].6'; 1735 '~S001R14 Auto Tip Changer Low 2 WB2[54].7'; 1736 '~S001R14 Auto Tip Changer Empty 2 WB2[54].8'; 1737 '~S001R14 Tip Wear Ratio Warning 2 - Touch Up Tip Dress Program WB2[54].9'; 1738 '~S001R14 Stud Weld 2 Maintenance Reqd WB2[54].10'; 1739 '~S001R14 Stud Weld 2 Low Stud Warning WB2[54].11'; 1740 '~Spare WB2[54].12'; 1741 '~S001R14 Rivet 2 Low Rivet Warning WB2[54].13'; 1742 '~S001R14 Rivet 2 - Skip Once Initiated from Robot TP WB2[54].14'; 1743 '~S001R14 Rivet 2 - Skip Remaining Initiated from Robot TP WB2[54].15'; 1744 '~S001R14 Rivet 2 Preventive Maintenace Required WB2[54].16'; 1745 '~S001R14 Rivet 2 Magazine Low WB2[54].17'; 1746 '~S001R14 Tip Change 2 Bypassed WB2[54].18'; 1747 '~S001R14 Laser Dirty Glass Warning WB2[54].19'; 1748 '~S001R14 Weld Ctrlr 2 Adaptive Mode Is Disabled WB2[54].20'; 1749 '~S001R14 Tip Cutter 2 Warning WB2[54].21'; 1750 '~S001R14 Rivet 2 Tape-Cut Required WB2[54].22'; 1751 '~S001R14 Mig Tip Nozzel Replacement Warning WB2[54].23'; 1752 '~S001R14 Mig Tip Nozzel Replacement Required WB2[54].24'; 1753 '~S001R14 Sealer Ctrlr 2 Minor Fault WB2[54].25'; 1754 '~S001R14 Sealer Ctrlr 2 Required Rezeroing WB2[54].26'; 1755 '~S001R14 Mig Barrel Replacement Warning WB2[54].27'; 1756 '~S001R14 Mig Barrel Replacement Required WB2[54].28'; 1757 '~S001R14 In Touch Up Mode WB2[54].29'; 1758 '~S001R14 Touch Up Mode Not Enabled WB2[54].30'; 1759 '~Spare WB2[54].31'; 1760 '~S001R14 Laser Controller Fault WB2[55].0'; 1761 '~S001R14 Laser Dirty Glass Warning WB2[55].1'; 1762 '~S001R14 Laser Warning WB2[55].2'; 1763 '~Spare WB2[55].3'; 1764 '~Spare WB2[55].4'; 1765 '~Spare WB2[55].5'; 1766 '~Spare WB2[55].6'; 1767 '~Spare WB2[55].7'; 1768 '~Spare WB2[55].8'; 1769 '~Spare WB2[55].9'; 1770 '~Spare WB2[55].10'; 1771 '~Spare WB2[55].11'; 1772 '~Spare WB2[55].12'; 1773 '~Spare WB2[55].13'; 1774 '~Spare WB2[55].14'; 1775 '~Spare WB2[55].15'; 1776 '~Spare WB2[55].16'; 1777 '~Spare WB2[55].17'; 1778 '~Spare WB2[55].18'; 1779 '~Spare WB2[55].19'; 1780 '~Spare WB2[55].20'; 1781 '~Spare WB2[55].21'; 1782 '~Spare WB2[55].22'; 1783 '~Spare WB2[55].23'; 1784 '~Spare WB2[55].24'; 1785 '~Spare WB2[55].25'; 1786 '~Spare WB2[55].26'; 1787 '~Spare WB2[55].27'; 1788 '~Spare WB2[55].28'; 1789 '~Spare WB2[55].29'; 1790 '~Spare WB2[55].30'; 1791 '~Spare WB2[55].31'; 1792 '~Spare WB2[56].0'; 1793 '~Spare WB2[56].1'; 1794 '~Spare WB2[56].2'; 1795 '~Spare WB2[56].3'; 1796 '~Spare WB2[56].4'; 1797 '~Spare WB2[56].5'; 1798 '~Spare WB2[56].6'; 1799 '~Spare WB2[56].7'; 1800 '~Spare WB2[56].8'; 1801 '~Spare WB2[56].9'; 1802 '~Spare WB2[56].10'; 1803 '~Spare WB2[56].11'; 1804 '~Spare WB2[56].12'; 1805 '~Spare WB2[56].13'; 1806 '~Spare WB2[56].14'; 1807 '~Spare WB2[56].15'; 1808 '~Spare WB2[56].16'; 1809 '~Spare WB2[56].17'; 1810 '~Spare WB2[56].18'; 1811 '~Spare WB2[56].19'; 1812 '~Spare WB2[56].20'; 1813 '~Spare WB2[56].21'; 1814 '~Spare WB2[56].22'; 1815 '~Spare WB2[56].23'; 1816 '~Spare WB2[56].24'; 1817 '~Spare WB2[56].25'; 1818 '~Spare WB2[56].26'; 1819 '~Spare WB2[56].27'; 1820 '~Spare WB2[56].28'; 1821 '~Spare WB2[56].29'; 1822 '~Spare WB2[56].30'; 1823 '~Spare WB2[56].31'; 1824 '~Spare WB2[57].0'; 1825 '~Spare WB2[57].1'; 1826 '~Spare WB2[57].2'; 1827 '~Spare WB2[57].3'; 1828 '~Spare WB2[57].4'; 1829 '~Spare WB2[57].5'; 1830 '~Spare WB2[57].6'; 1831 '~Spare WB2[57].7'; 1832 '~Spare WB2[57].8'; 1833 '~Spare WB2[57].9'; 1834 '~Spare WB2[57].10'; 1835 '~Spare WB2[57].11'; 1836 '~Spare WB2[57].12'; 1837 '~Spare WB2[57].13'; 1838 '~Spare WB2[57].14'; 1839 '~Spare WB2[57].15'; 1840 '~Spare WB2[57].16'; 1841 '~Spare WB2[57].17'; 1842 '~Spare WB2[57].18'; 1843 '~Spare WB2[57].19'; 1844 '~Spare WB2[57].20'; 1845 '~Spare WB2[57].21'; 1846 '~Spare WB2[57].22'; 1847 '~Spare WB2[57].23'; 1848 '~Spare WB2[57].24'; 1849 '~Spare WB2[57].25'; 1850 '~Spare WB2[57].26'; 1851 '~Spare WB2[57].27'; 1852 '~Spare WB2[57].28'; 1853 '~Spare WB2[57].29'; 1854 '~Spare WB2[57].30'; 1855 '~Spare WB2[57].31'; 1856 '~S001R15 Waiting Zone #1 Not Clear WB2[58].0'; 1857 '~S001R15 Waiting Zone #2 Not Clear WB2[58].1'; 1858 '~S001R15 Waiting Zone #3 Not Clear WB2[58].2'; 1859 '~S001R15 Waiting Zone #4 Not Clear WB2[58].3'; 1860 '~S001R15 Waiting Zone #5 Not Clear WB2[58].4'; 1861 '~S001R15 Waiting Zone #6 Not Clear WB2[58].5'; 1862 '~S001R15 Waiting Zone #7 Not Clear WB2[58].6'; 1863 '~S001R15 Waiting Zone #8 Not Clear WB2[58].7'; 1864 '~S001R15 Waiting Zone #9 Not Clear WB2[58].8'; 1865 '~S001R15 Waiting Zone #10 Not Clear WB2[58].9'; 1866 '~S001R15 Waiting Zone #11 Not Clear WB2[58].10'; 1867 '~S001R15 Waiting Zone #12 Not Clear WB2[58].11'; 1868 '~S001R15 Waiting Zone #13 Not Clear WB2[58].12'; 1869 '~S001R15 Waiting Zone #14 Not Clear WB2[58].13'; 1870 '~S001R15 Waiting Tip Dress Zone #1 Not Clear WB2[58].14'; 1871 '~S001R15 Waiting Tip Dress Zone #2 Not Clear WB2[58].15'; 1872 '~S001R15 Adjacent Robot xx-xx In Teach WB2[58].16'; 1873 '~S001R15 Adjacent Robot xx-xx In Teach WB2[58].17'; 1874 '~S001R15 Adjacent Robot xx-xx In Teach WB2[58].18'; 1875 '~S001R15 Adjacent Robot xx-xx In Teach WB2[58].19'; 1876 '~S001R15 Adjacent Robot xx-xx In Teach WB2[58].20'; 1877 '~S001R15 Adjacent Robot xx-xx In Teach WB2[58].21'; 1878 '~S001R15 Adjacent Robot xx-xx In Teach WB2[58].22'; 1879 '~S001R15 Adjacent Robot xx-xx In Teach WB2[58].23'; 1880 '~S001R15 Adjacent Robot xx-xx In Teach WB2[58].24'; 1881 '~S001R15 Adjacent Robot xx-xx In Teach WB2[58].25'; 1882 '~Spare WB2[58].26'; 1883 '~Spare WB2[58].27'; 1884 '~Spare WB2[58].28'; 1885 '~S001R15 Robot Not Clear Of Fixture WB2[58].29'; 1886 '~Spare WB2[58].30'; 1887 '~Spare WB2[58].31'; 1888 '~Spare WB2[59].0'; 1889 '~Spare WB2[59].1'; 1890 '~Spare WB2[59].2'; 1891 '~Spare WB2[59].3'; 1892 '~Spare WB2[59].4'; 1893 '~Spare WB2[59].5'; 1894 '~Spare WB2[59].6'; 1895 '~Spare WB2[59].7'; 1896 '~Spare WB2[59].8'; 1897 '~Spare WB2[59].9'; 1898 '~Spare WB2[59].10'; 1899 '~Spare WB2[59].11'; 1900 '~Spare WB2[59].12'; 1901 '~Spare WB2[59].13'; 1902 '~Spare WB2[59].14'; 1903 '~Spare WB2[59].15'; 1904 '~Spare WB2[59].16'; 1905 '~Spare WB2[59].17'; 1906 '~Spare WB2[59].18'; 1907 '~Spare WB2[59].19'; 1908 '~Spare WB2[59].20'; 1909 '~Spare WB2[59].21'; 1910 '~Spare WB2[59].22'; 1911 '~Spare WB2[59].23'; 1912 '~Spare WB2[59].24'; 1913 '~Spare WB2[59].25'; 1914 '~Spare WB2[59].26'; 1915 '~Spare WB2[59].27'; 1916 '~Spare WB2[59].28'; 1917 '~Spare WB2[59].29'; 1918 '~Spare WB2[59].30'; 1919 '~Spare WB2[59].31'; 1920 '~S001R15 Cycle Overtime WB2[60].0'; 1921 '~S001R15 In Bypass WB2[60].1'; 1922 '~S001R15 Battery Low WB2[60].2'; 1923 '~S001R15 Servo Over Torque WB2[60].3'; 1924 '~S001R15 Process Retry In Progress WB2[60].4'; 1925 '~Spare WB2[60].5'; 1926 '~S001R15 Robot Edit Occurred Ext App WB2[60].6'; 1927 '~S001R15 Robot Input Simmed WB2[60].7'; 1928 '~S001R15 Robot Output Simmed WB2[60].8'; 1929 '~Spare WB2[60].9'; 1930 '~Spare WB2[60].10'; 1931 '~Spare WB2[60].11'; 1932 '~Spare WB2[60].12'; 1933 '~Spare WB2[60].13'; 1934 '~Spare WB2[60].14'; 1935 '~Spare WB2[60].15'; 1936 '~S001R15F1B1.M.ModuleFlt - Externa App 1 I/O Module Warning WB2[60].16'; 1937 '~S001R15F2B1.M.ModuleFlt - Externa App 2 I/O Module Warning WB2[60].17'; 1938 '~S001R15F3B1.M.ModuleFlt - Externa App 3 I/O Module Warning WB2[60].18'; 1939 '~Spare WB2[60].19'; 1940 '~Spare WB2[60].20'; 1941 '~Spare WB2[60].21'; 1942 '~Spare WB2[60].22'; 1943 '~Spare WB2[60].23'; 1944 '~S001R15ES1 - S001R15 EtherNet Switch Port At Half Duplex WB2[60].24'; 1945 '~S001R15ES1 - S001R15 EtherNet Switch Config Changes Not Saved WB2[60].25'; 1946 '~S001R15ES1 - S001R15 EtherNet Switch Configuration Changed WB2[60].26'; 1947 '~S001R15ES1 - S001R15 EtherNet Switch Port With Excessive Errors WB2[60].27'; 1948 '~S001R15ES1 - S001R15 EtherNet Switch Port With Utilization Warning WB2[60].28'; 1949 '~S001R15ES1 - S001R15 EtherNet Switch Changes Require Reboot WB2[60].29'; 1950 '~Spare WB2[60].30'; 1951 '~Spare WB2[60].31'; 1952 '~Spare WB2[61].0'; 1953 '~Spare WB2[61].1'; 1954 '~S001R15 Servo Gun Tip Calib Request 1 WB2[61].2'; 1955 '~S001R15 I-Available Warning 1 WB2[61].3'; 1956 '~S001R15 Tip Dress Motor 1 Fault Bypassed WB2[61].4'; 1957 '~S001R15 Tip Change Notice 1 WB2[61].5'; 1958 '~S001R15 Bypass Tip Dresser 1 Selected WB2[61].6'; 1959 '~S001R15 Auto Tip Changer Low 1 WB2[61].7'; 1960 '~S001R15 Auto Tip Changer Empty 1 WB2[61].8'; 1961 '~S001R15 Tip Wear Ratio Warning 1 - Touch Up Tip Dress Program WB2[61].9'; 1962 '~S001R15 Stud Weld 1 Maintenance Reqd WB2[61].10'; 1963 '~S001R15 Stud Weld 1 Low Stud Warning WB2[61].11'; 1964 '~Spare WB2[61].12'; 1965 '~S001R15 Rivet 1 Low Rivet Warning WB2[61].13'; 1966 '~S001R15 Rivet 1 - Skip Once Initiated from Robot TP WB2[61].14'; 1967 '~S001R15 Rivet 1 - Skip Remaining Initiated from Robot TP WB2[61].15'; 1968 '~S001R15 Rivet 1 Preventive Maintenace Required WB2[61].16'; 1969 '~S001R15 Rivet 1 Magazine Low WB2[61].17'; 1970 '~S001R15 Tip Change 1 Bypassed WB2[61].18'; 1971 '~S001R15 Mig Weld Fluid Level Low WB2[61].19'; 1972 '~S001R15 Weld Ctrlr 1 Adaptive Mode Is Disabled WB2[61].20'; 1973 '~S001R15 Tip Cutter 1 Warning WB2[61].21'; 1974 '~S001R15 Rivet 1 Tape-Cut Required WB2[61].22'; 1975 '~S001R15 Wire Feeder Motor Over Current WB2[61].23'; 1976 '~Spare WB2[61].24'; 1977 '~S001R15 Sealer Ctrlr 1 Minor Fault WB2[61].25'; 1978 '~S001R15 Sealer Ctrlr 1 Required Rezeroing WB2[61].26'; 1979 '~S001R15 Loaded To Average WB2[61].27'; 1980 '~S001R15 Vision Process Aborted WB2[61].28'; 1981 '~S001R15 Vision System Trending WB2[61].29'; 1982 '~S001R15 Vision Out Of Tolerance WB2[61].30'; 1983 '~Spare WB2[61].31'; 1984 '~Spare WB2[62].0'; 1985 '~Spare WB2[62].1'; 1986 '~S001R15 Servo Gun Tip Calib Request 2 WB2[62].2'; 1987 '~S001R15 I-Available Warning 2 WB2[62].3'; 1988 '~S001R15 Tip Dress Motor 2 Fault Bypassed WB2[62].4'; 1989 '~S001R15 Tip Change Notice 2 WB2[62].5'; 1990 '~S001R15 Bypass Tip Dresser 2 Selected WB2[62].6'; 1991 '~S001R15 Auto Tip Changer Low 2 WB2[62].7'; 1992 '~S001R15 Auto Tip Changer Empty 2 WB2[62].8'; 1993 '~S001R15 Tip Wear Ratio Warning 2 - Touch Up Tip Dress Program WB2[62].9'; 1994 '~S001R15 Stud Weld 2 Maintenance Reqd WB2[62].10'; 1995 '~S001R15 Stud Weld 2 Low Stud Warning WB2[62].11'; 1996 '~Spare WB2[62].12'; 1997 '~S001R15 Rivet 2 Low Rivet Warning WB2[62].13'; 1998 '~S001R15 Rivet 2 - Skip Once Initiated from Robot TP WB2[62].14'; 1999 '~S001R15 Rivet 2 - Skip Remaining Initiated from Robot TP WB2[62].15'; 2000 '~S001R15 Rivet 2 Preventive Maintenace Required WB2[62].16'; 2001 '~S001R15 Rivet 2 Magazine Low WB2[62].17'; 2002 '~S001R15 Tip Change 2 Bypassed WB2[62].18'; 2003 '~S001R15 Laser Dirty Glass Warning WB2[62].19'; 2004 '~S001R15 Weld Ctrlr 2 Adaptive Mode Is Disabled WB2[62].20'; 2005 '~S001R15 Tip Cutter 2 Warning WB2[62].21'; 2006 '~S001R15 Rivet 2 Tape-Cut Required WB2[62].22'; 2007 '~S001R15 Mig Tip Nozzel Replacement Warning WB2[62].23'; 2008 '~S001R15 Mig Tip Nozzel Replacement Required WB2[62].24'; 2009 '~S001R15 Sealer Ctrlr 2 Minor Fault WB2[62].25'; 2010 '~S001R15 Sealer Ctrlr 2 Required Rezeroing WB2[62].26'; 2011 '~S001R15 Mig Barrel Replacement Warning WB2[62].27'; 2012 '~S001R15 Mig Barrel Replacement Required WB2[62].28'; 2013 '~S001R15 In Touch Up Mode WB2[62].29'; 2014 '~S001R15 Touch Up Mode Not Enabled WB2[62].30'; 2015 '~Spare WB2[62].31'; 2016 '~S001R15 Laser Controller Fault WB2[63].0'; 2017 '~S001R15 Laser Dirty Glass Warning WB2[63].1'; 2018 '~S001R15 Laser Warning WB2[63].2'; 2019 '~Spare WB2[63].3'; 2020 '~Spare WB2[63].4'; 2021 '~Spare WB2[63].5'; 2022 '~Spare WB2[63].6';